// TIA Portal project "Motor with VFD+PID" (V20)

(* hardware
DEVICE "S7-1200 station_1"  S7-1200 Station
   slot 0: "Rack_0"  S7-1200 Rack  Rack  V1.0
   slot 1: "PLC_1"  CPU 1214C DC/DC/DC  6ES7 214-1AG40-0XB0  V4.7
DEVICE "HMI_1"  KTP700 Basic PN
   slot 0: "HMI_1"  KTP700 Basic PN  6AV2 123-2GB03-0AX0  17.0.0.0
   slot 1: "HMI_RT_1"  KTP700 Basic PN  6AV2 123-2GB03-0AX0  17.0.0.0
   slot 5: "HMI_1.IE_CP_1"  PROFINET Interface  17.0.0.0
      slot 1: "PROFINET Interface_1"  PROFINET Interface
         slot 1: "Port_1"  Port
*)

// ===== PLC "PLC_1"  CPU 1214C DC/DC/DC =====

VAR_GLOBAL   // PLC tag table "Default tag table"
   "Start_PB" AT %I0.0 : Bool;
   "Stop_PB" AT %I0.1 : Bool;
   "VFD_Fault" AT %I0.2 : Bool;
   "VFD_Running_FB" AT %I0.3 : Bool;
   "Reset_PB" AT %I0.4 : Bool;
   "VFD_Run_CMD" AT %Q0.0 : Bool;
   "VFD_Reset_CMD" AT %Q0.1 : Bool;
   "Motor_Run_Latch" AT %M0.0 : Bool;
   "Alarm_Active" AT %M0.1 : Bool;
   "Auto_Mode" AT %M0.2 : Bool;
   "Manual_Mode" AT %M0.3 : Bool;
   "HMI_START" AT %M0.4 : Bool;
   "HMI_STOP" AT %M0.5 : Bool;
   "HMI_RESET" AT %M0.6 : Bool;
END_VAR

DATA_BLOCK "DB_VFD_Motor"   // DB1
{ S7_Optimized_Access := 'TRUE' }
VERSION : 0.1
   VAR RETAIN
      Speed_setpoint_hz : Real := 25.0;
   END_VAR
   VAR
      Max_Hz : Real := 50.0;
      Min_Hz : Real;
      Pressure_Setpoint : Real := 6.0;
      Ramp_Output : Real;
      Ramp_Step : Real := 1.0;
      Pressure_Actual : Real := 4.0;
      PID_Error : Real;
   END_VAR
   VAR RETAIN
      Ramp_time : Real;
   END_VAR
   VAR
      Low_Pressure_timer_Done : Bool;
      Min_Pressure_Limit : Real := 1.0;
      Max_Pressure_Limit : Real := 8.0;
      Manual_Speed_Hz : Real := 20.0;
      Overpressure_Alarm : Bool;
      Low_Pressure_Alarm : Bool;
      Fault_code : Int;
      Actual_speed_hz : Real;
      Output_scaled : Int;
   END_VAR
BEGIN
END_DATA_BLOCK

// folder: System blocks/Program resources

DATA_BLOCK "TON"   // DB2
{ S7_Optimized_Access := 'TRUE' }
AUTHOR : Simatic
FAMILY : IEC
NAME : IEC_TMR
VERSION : 1.0
// stored: InstanceOfName IEC_TIMER
"IEC_TIMER"
BEGIN
END_DATA_BLOCK

// folder: (top level)

ORGANIZATION_BLOCK "Main"   // OB1, LAD, ProgramCycle
TITLE = "Main Program Sweep (Cycle)"
{ S7_Optimized_Access := 'TRUE' }
VERSION : 0.1
   VAR_INPUT
      Initial_Call : Bool;   // Initial call of this OB
      Remanence : Bool;   // =True, if remanent data are available
   END_VAR
BEGIN

REGION Network 1: Start/Stop Safety Logic
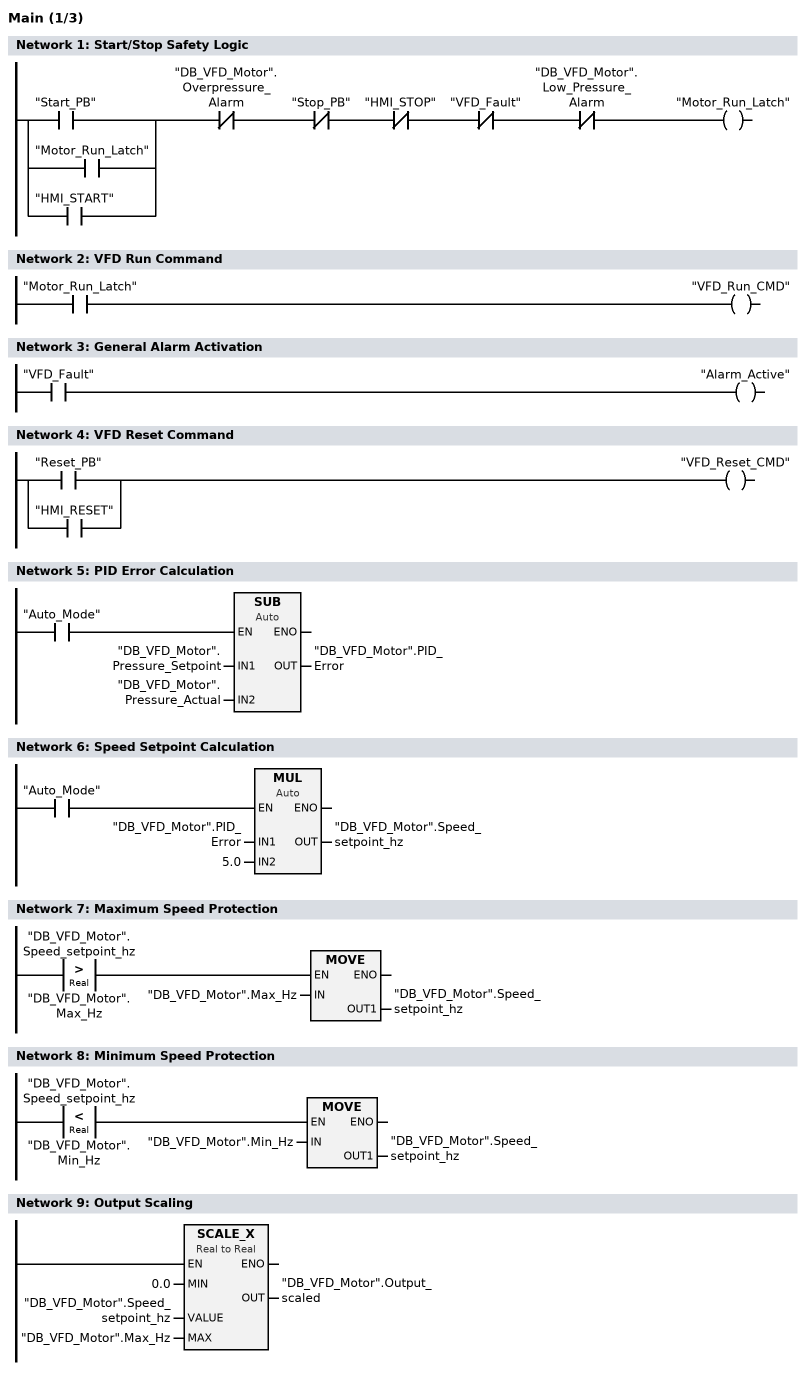
   RUNG wire#powerrail
      Contact( "Start_PB" )
      wire#w1
      I_Contact( "DB_VFD_Motor".Overpressure_Alarm )
      I_Contact( "Stop_PB" )
      I_Contact( "HMI_STOP" )
      I_Contact( "VFD_Fault" )
      I_Contact( "DB_VFD_Motor".Low_Pressure_Alarm )
      Coil( "Motor_Run_Latch" )
   END_RUNG
   RUNG wire#powerrail
      Contact( "Motor_Run_Latch" )
   END_RUNG wire#w1
   RUNG wire#powerrail
      Contact( "HMI_START" )
   END_RUNG wire#w1
   // the same network as SCL:
   "Motor_Run_Latch" := ("Start_PB" OR "Motor_Run_Latch" OR "HMI_START") AND NOT "DB_VFD_Motor".Overpressure_Alarm AND NOT "Stop_PB" AND NOT "HMI_STOP" AND NOT "VFD_Fault" AND NOT "DB_VFD_Motor".Low_Pressure_Alarm;
END_REGION

REGION Network 2: VFD Run Command
   RUNG wire#powerrail
      Contact( "Motor_Run_Latch" )
      Coil( "VFD_Run_CMD" )
   END_RUNG
   // the same network as SCL:
   "VFD_Run_CMD" := "Motor_Run_Latch";
END_REGION

REGION Network 3: General Alarm Activation
   RUNG wire#powerrail
      Contact( "VFD_Fault" )
      Coil( "Alarm_Active" )
   END_RUNG
   // the same network as SCL:
   "Alarm_Active" := "VFD_Fault";
END_REGION

REGION Network 4: VFD Reset Command
   RUNG wire#powerrail
      Contact( "Reset_PB" )
      wire#w1
      Coil( "VFD_Reset_CMD" )
   END_RUNG
   RUNG wire#powerrail
      Contact( "HMI_RESET" )
   END_RUNG wire#w1
   // the same network as SCL:
   "VFD_Reset_CMD" := "Reset_PB" OR "HMI_RESET";
END_REGION

REGION Network 5: PID Error Calculation
   RUNG wire#powerrail
      Contact( "Auto_Mode" )
      Sub(in1 := "DB_VFD_Motor".Pressure_Setpoint, in2 := "DB_VFD_Motor".Pressure_Actual, out => "DB_VFD_Motor".PID_Error)
   END_RUNG
   // the same network as SCL:
   IF "Auto_Mode" THEN
       "DB_VFD_Motor".PID_Error := "DB_VFD_Motor".Pressure_Setpoint - "DB_VFD_Motor".Pressure_Actual;
   END_IF;
END_REGION

REGION Network 6: Speed Setpoint Calculation
   RUNG wire#powerrail
      Contact( "Auto_Mode" )
      Mul(in1 := "DB_VFD_Motor".PID_Error, in2 := 5.0, out => "DB_VFD_Motor".Speed_setpoint_hz)
   END_RUNG
   // the same network as SCL:
   IF "Auto_Mode" THEN "DB_VFD_Motor".Speed_setpoint_hz := "DB_VFD_Motor".PID_Error * 5.0; END_IF;
END_REGION

REGION Network 7: Maximum Speed Protection
   RUNG wire#powerrail
      { S7_Templates := "SrcType := Real" } GT_Contact(in1 := "DB_VFD_Motor".Speed_setpoint_hz, in2 := "DB_VFD_Motor".Max_Hz)
      Move(in := "DB_VFD_Motor".Max_Hz, out1 => "DB_VFD_Motor".Speed_setpoint_hz)
   END_RUNG
   // the same network as SCL:
   IF "DB_VFD_Motor".Speed_setpoint_hz > "DB_VFD_Motor".Max_Hz THEN
       "DB_VFD_Motor".Speed_setpoint_hz := "DB_VFD_Motor".Max_Hz;
   END_IF;
END_REGION

REGION Network 8: Minimum Speed Protection
   RUNG wire#powerrail
      { S7_Templates := "SrcType := Real" } LT_Contact(in1 := "DB_VFD_Motor".Speed_setpoint_hz, in2 := "DB_VFD_Motor".Min_Hz)
      Move(in := "DB_VFD_Motor".Min_Hz, out1 => "DB_VFD_Motor".Speed_setpoint_hz)
   END_RUNG
   // the same network as SCL:
   IF "DB_VFD_Motor".Speed_setpoint_hz < "DB_VFD_Motor".Min_Hz THEN
       "DB_VFD_Motor".Speed_setpoint_hz := "DB_VFD_Motor".Min_Hz;
   END_IF;
END_REGION

REGION Network 9: Output Scaling
   RUNG wire#powerrail
      { S7_Templates := "[SrcType := Real, DestType := Real]" } Scale(min := 0.0, value := "DB_VFD_Motor".Speed_setpoint_hz, max := "DB_VFD_Motor".Max_Hz, out => "DB_VFD_Motor".Output_scaled)
   END_RUNG
   // the same network as SCL:
   "DB_VFD_Motor".Output_scaled := SCALE_X(MIN := 0.0, VALUE := "DB_VFD_Motor".Speed_setpoint_hz, MAX := "DB_VFD_Motor".Max_Hz);
END_REGION

REGION Network 10: Motor Speed Update
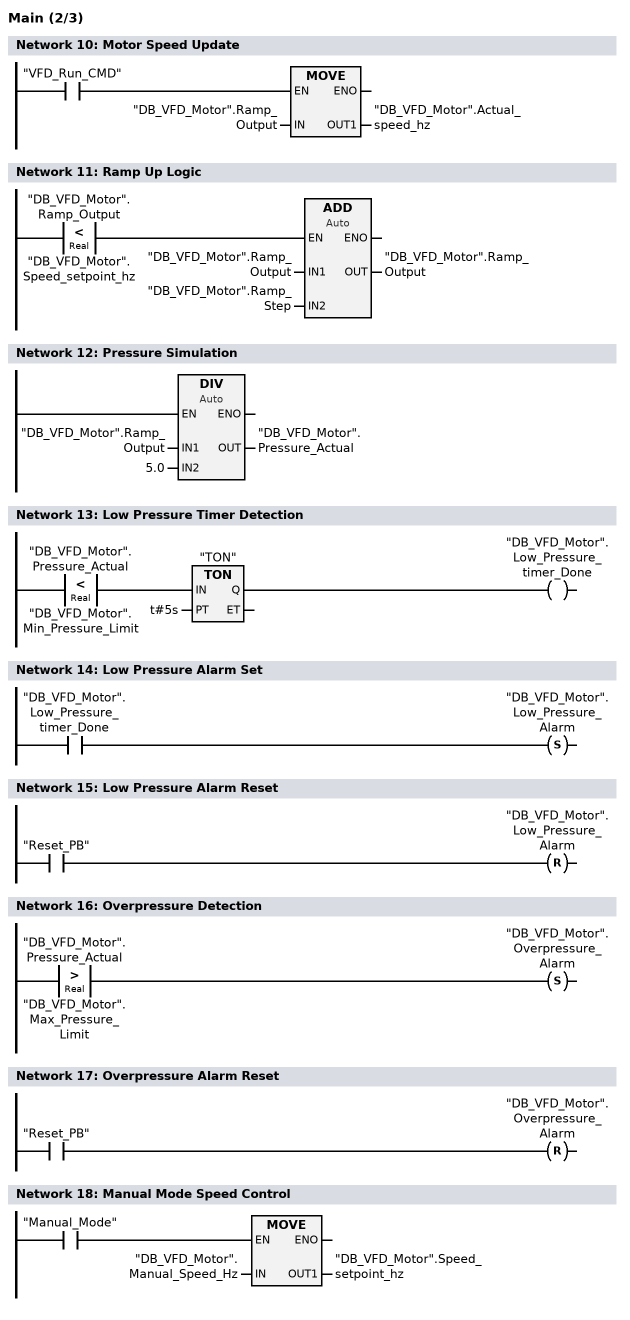
   RUNG wire#powerrail
      Contact( "VFD_Run_CMD" )
      Move(in := "DB_VFD_Motor".Ramp_Output, out1 => "DB_VFD_Motor".Actual_speed_hz)
   END_RUNG
   // the same network as SCL:
   IF "VFD_Run_CMD" THEN "DB_VFD_Motor".Actual_speed_hz := "DB_VFD_Motor".Ramp_Output; END_IF;
END_REGION

REGION Network 11: Ramp Up Logic
   RUNG wire#powerrail
      { S7_Templates := "SrcType := Real" } LT_Contact(in1 := "DB_VFD_Motor".Ramp_Output, in2 := "DB_VFD_Motor".Speed_setpoint_hz)
      Add(in1 := "DB_VFD_Motor".Ramp_Output, in2 := "DB_VFD_Motor".Ramp_Step, out => "DB_VFD_Motor".Ramp_Output)
   END_RUNG
   // the same network as SCL:
   IF "DB_VFD_Motor".Ramp_Output < "DB_VFD_Motor".Speed_setpoint_hz THEN
       "DB_VFD_Motor".Ramp_Output := "DB_VFD_Motor".Ramp_Output + "DB_VFD_Motor".Ramp_Step;
   END_IF;
END_REGION

REGION Network 12: Pressure Simulation
   RUNG wire#powerrail
      Div(in1 := "DB_VFD_Motor".Ramp_Output, in2 := 5.0, out => "DB_VFD_Motor".Pressure_Actual)
   END_RUNG
   // the same network as SCL:
   "DB_VFD_Motor".Pressure_Actual := "DB_VFD_Motor".Ramp_Output / 5.0;
END_REGION

REGION Network 13: Low Pressure Timer Detection
   "TON".TON(IN := "DB_VFD_Motor".Pressure_Actual < "DB_VFD_Motor".Min_Pressure_Limit, PT := t#5s);
   "DB_VFD_Motor".Low_Pressure_timer_Done := "TON".Q;
END_REGION

REGION Network 14: Low Pressure Alarm Set
   RUNG wire#powerrail
      Contact( "DB_VFD_Motor".Low_Pressure_timer_Done )
      S_Coil( "DB_VFD_Motor".Low_Pressure_Alarm )
   END_RUNG
   // the same network as SCL:
   IF "DB_VFD_Motor".Low_Pressure_timer_Done THEN "DB_VFD_Motor".Low_Pressure_Alarm := TRUE; END_IF;
END_REGION

REGION Network 15: Low Pressure Alarm Reset
   RUNG wire#powerrail
      Contact( "Reset_PB" )
      R_Coil( "DB_VFD_Motor".Low_Pressure_Alarm )
   END_RUNG
   // the same network as SCL:
   IF "Reset_PB" THEN "DB_VFD_Motor".Low_Pressure_Alarm := FALSE; END_IF;
END_REGION

REGION Network 16: Overpressure Detection
   RUNG wire#powerrail
      { S7_Templates := "SrcType := Real" } GT_Contact(in1 := "DB_VFD_Motor".Pressure_Actual, in2 := "DB_VFD_Motor".Max_Pressure_Limit)
      S_Coil( "DB_VFD_Motor".Overpressure_Alarm )
   END_RUNG
   // the same network as SCL:
   IF "DB_VFD_Motor".Pressure_Actual > "DB_VFD_Motor".Max_Pressure_Limit THEN
       "DB_VFD_Motor".Overpressure_Alarm := TRUE;
   END_IF;
END_REGION

REGION Network 17: Overpressure Alarm Reset
   RUNG wire#powerrail
      Contact( "Reset_PB" )
      R_Coil( "DB_VFD_Motor".Overpressure_Alarm )
   END_RUNG
   // the same network as SCL:
   IF "Reset_PB" THEN "DB_VFD_Motor".Overpressure_Alarm := FALSE; END_IF;
END_REGION

REGION Network 18: Manual Mode Speed Control
   RUNG wire#powerrail
      Contact( "Manual_Mode" )
      Move(in := "DB_VFD_Motor".Manual_Speed_Hz, out1 => "DB_VFD_Motor".Speed_setpoint_hz)
   END_RUNG
   // the same network as SCL:
   IF "Manual_Mode" THEN "DB_VFD_Motor".Speed_setpoint_hz := "DB_VFD_Motor".Manual_Speed_Hz; END_IF;
END_REGION

REGION Network 19: VFD Fault Code Assignment
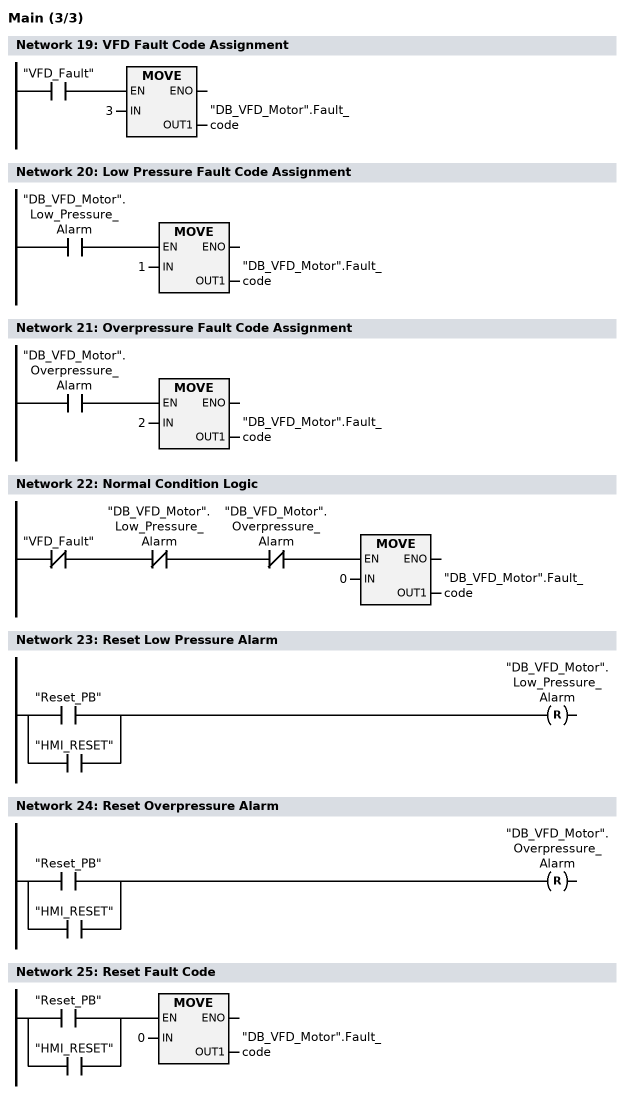
   RUNG wire#powerrail
      Contact( "VFD_Fault" )
      Move(in := 3, out1 => "DB_VFD_Motor".Fault_code)
   END_RUNG
   // the same network as SCL:
   IF "VFD_Fault" THEN "DB_VFD_Motor".Fault_code := 3; END_IF;
END_REGION

REGION Network 20: Low Pressure Fault Code Assignment
   RUNG wire#powerrail
      Contact( "DB_VFD_Motor".Low_Pressure_Alarm )
      Move(in := 1, out1 => "DB_VFD_Motor".Fault_code)
   END_RUNG
   // the same network as SCL:
   IF "DB_VFD_Motor".Low_Pressure_Alarm THEN "DB_VFD_Motor".Fault_code := 1; END_IF;
END_REGION

REGION Network 21: Overpressure Fault Code Assignment
   RUNG wire#powerrail
      Contact( "DB_VFD_Motor".Overpressure_Alarm )
      Move(in := 2, out1 => "DB_VFD_Motor".Fault_code)
   END_RUNG
   // the same network as SCL:
   IF "DB_VFD_Motor".Overpressure_Alarm THEN "DB_VFD_Motor".Fault_code := 2; END_IF;
END_REGION

REGION Network 22: Normal Condition Logic
   RUNG wire#powerrail
      I_Contact( "VFD_Fault" )
      I_Contact( "DB_VFD_Motor".Low_Pressure_Alarm )
      I_Contact( "DB_VFD_Motor".Overpressure_Alarm )
      Move(in := 0, out1 => "DB_VFD_Motor".Fault_code)
   END_RUNG
   // the same network as SCL:
   IF NOT "VFD_Fault" AND NOT "DB_VFD_Motor".Low_Pressure_Alarm AND NOT "DB_VFD_Motor".Overpressure_Alarm THEN
       "DB_VFD_Motor".Fault_code := 0;
   END_IF;
END_REGION

REGION Network 23: Reset Low Pressure Alarm
   RUNG wire#powerrail
      Contact( "Reset_PB" )
      wire#w1
      R_Coil( "DB_VFD_Motor".Low_Pressure_Alarm )
   END_RUNG
   RUNG wire#powerrail
      Contact( "HMI_RESET" )
   END_RUNG wire#w1
   // the same network as SCL:
   IF "Reset_PB" OR "HMI_RESET" THEN "DB_VFD_Motor".Low_Pressure_Alarm := FALSE; END_IF;
END_REGION

REGION Network 24: Reset Overpressure Alarm
   RUNG wire#powerrail
      Contact( "Reset_PB" )
      wire#w1
      R_Coil( "DB_VFD_Motor".Overpressure_Alarm )
   END_RUNG
   RUNG wire#powerrail
      Contact( "HMI_RESET" )
   END_RUNG wire#w1
   // the same network as SCL:
   IF "Reset_PB" OR "HMI_RESET" THEN "DB_VFD_Motor".Overpressure_Alarm := FALSE; END_IF;
END_REGION

REGION Network 25: Reset Fault Code
   RUNG wire#powerrail
      Contact( "Reset_PB" )
      wire#w1
      Move(in := 0, out1 => "DB_VFD_Motor".Fault_code)
   END_RUNG
   RUNG wire#powerrail
      Contact( "HMI_RESET" )
   END_RUNG wire#w1
   // the same network as SCL:
   IF "Reset_PB" OR "HMI_RESET" THEN "DB_VFD_Motor".Fault_code := 0; END_IF;
END_REGION
END_ORGANIZATION_BLOCK

(* ===== HMI "HMI_RT_1" =====
system functions are stored by id; their names below are inferred from use
connection "HMI_Connection_1": ETHERNET, SMART_S7_1200_OMS

HMI tags "Default tag table"
   "Tag_ScreenNumber" : UInt, internal
   "Motor_Run_Latch" : Bool = PLC Motor_Run_Latch AT %M0.0, 1 s
   "Alarm_Active" : Bool = PLC Alarm_Active AT %M0.1, 1 s
   "Auto_Mode" : Bool = PLC Auto_Mode AT %M0.2, 1 s
   "Manual_Mode" : Bool = PLC Manual_Mode AT %M0.3, 1 s
   "HMI_START" : Bool = PLC HMI_START AT %M0.4, 1 s
   "HMI_STOP" : Bool = PLC HMI_STOP AT %M0.5, 1 s
   "HMI_RESET" : Bool = PLC HMI_RESET AT %M0.6, 1 s
   "DB_VFD_Motor_Pressure_Setpoint" : Real = PLC DB_VFD_Motor.Pressure_Setpoint, 1 s
   "DB_VFD_Motor_Pressure_Actual" : Real = PLC DB_VFD_Motor.Pressure_Actual, 1 s
   "DB_VFD_Motor_Actual_speed_hz" : Real = PLC DB_VFD_Motor.Actual_speed_hz, 1 s
   "DB_VFD_Motor_Output_scaled" : Int = PLC DB_VFD_Motor.Output_scaled, 1 s
   "DB_VFD_Motor_Manual_Speed_Hz" : Real = PLC DB_VFD_Motor.Manual_Speed_Hz, 1 s
   "DB_VFD_Motor_PID_Error" : Real = PLC DB_VFD_Motor.PID_Error, 1 s
   "DB_VFD_Motor_Speed_setpoint_hz" : Real = PLC DB_VFD_Motor.Speed_setpoint_hz, 1 s
   "DB_VFD_Motor_Ramp_Output" : Real = PLC DB_VFD_Motor.Ramp_Output, 1 s
   "DB_VFD_Motor_Min_Pressure_Limit" : Real = PLC DB_VFD_Motor.Min_Pressure_Limit, 1 s
   "DB_VFD_Motor_Max_Pressure_Limit" : Real = PLC DB_VFD_Motor.Max_Pressure_Limit, 1 s
   "DB_VFD_Motor_Ramp_Step" : Real = PLC DB_VFD_Motor.Ramp_Step, 1 s
   "DB_VFD_Motor_Fault_code" : Int = PLC DB_VFD_Motor.Fault_code, 1 s
   "VFD_Fault" : Bool = PLC VFD_Fault AT %I0.2, 1 s
   "DB_VFD_Motor_Low_Pressure_Alarm" : Bool = PLC DB_VFD_Motor.Low_Pressure_Alarm, 1 s
   "DB_VFD_Motor_Overpressure_Alarm" : Bool = PLC DB_VFD_Motor.Overpressure_Alarm, 1 s

text list "ACTIVE": 0 'INACTIVE'; 1 'ACTIVE'

text list "RUNNING": 0 'STOPPED'; 1 'RUNNING'

text list "ALARM": 0 'NO ALARM'; 1 'ALARM'

text list "NO FAULT": 0 'NO FAULT'; 1 'VFD FAULT ACTIVE'

text list "NO ALARM": 0 'NO ALARM'; 1 'LOW PRESSURE ACTIVE'

text list "OVERPRESSURE ACTIVE": 0 'NO ALARM'; 1 'OVERPRESSURE ACTIVE'

Template "Template_1" 800x480
   Button "Exit" at 714,429 size 71x50; TextOff 'Exit'; PictureOff "ExitRuntime_KTP700_Basic_PN_TR"; PictureOn "ExitRuntime_KTP700_Basic_PN_TR"
      on Release: StopRuntime(0)
   Button "Template_Button" at 614,429 size 71x50; TextOff 'Text'
   Button "Template_Button_1" at 514,429 size 71x50; TextOff 'Text'
   Button "Template_Button_2" at 414,429 size 71x50; TextOff 'Text'
   Button "Template_Button_3" at 314,429 size 71x50; TextOff 'Text'
   Button "Template_Button_4" at 214,429 size 71x50; TextOff 'Text'
   Button "Template_Button_5" at 114,429 size 71x50; TextOff 'Text'
   Button "Start screen" at 14,429 size 71x50; TextOff 'Start screen'; PictureOff "NavigateHome_KTP700_Basic_PN_TR"; PictureOn "NavigateHome_KTP700_Basic_PN_TR"
      on Release: ActivateScreen("Main Overview", 0)
   SymbolicIOField "Symbolic_IO_Field_Screen" at 93,9 size 600x33; TextOff '0'; TextOn '1'; TextList "TextList_ScreenNames"
      ProcessValue <- "Tag_ScreenNumber"
      on Change: ActivateScreenByNumber("Tag_ScreenNumber", 0)
   DateTimeField "HmiScreenItemData" at 695,25 size 105x25
   DateTimeField "HmiScreenItemData_1" at 695,0 size 105x25
   GraphicView "Logo" at 0,0 size 91x51; Picture "Logo of HMI_1"

screen "Main Overview" 800x480, template "Template_1"
   on GenerateScreen: SetTag("Tag_ScreenNumber", 1)
   GraphicView "Graphic view_1" at 2,1 size 796x478; Picture "ChatGPT Image 23 Ιουν 2026, 10_41_49 μ.μ."
   TextField "Text field_1" at 235,6 size 313x27; Text 'VFD PUMP PRESSURE CONTROL'
   GraphicView "Graphic view_2" at 123,75 size 264x225; Picture "ChatGPT Image 23 Ιουν 2026, 10_44_50 μ.μ."
   TextField "Text field_2" at 304,43 size 150x25; Text 'MAIN OVERVIEW'
   Button "Button_1" at 146,332 size 144x62; TextOff 'START'
      on Press: function_b14e0dd5("HMI_START", 0)
   Button "Button_2" at 1,414 size 194x65; TextOff 'HOME'
   Button "Button_3" at 195,414 size 204x65; TextOff 'CONTROL'
      on Press: ActivateScreen("Control", 0)
   Button "Button_4" at 398,414 size 200x65; TextOff 'ALARMS'
      on Press: ActivateScreen("Alarm Page", 0)
   Button "Button_5" at 597,414 size 200x65; TextOff 'DIAGNOSTICS'
      on Press: ActivateScreen("Diagnostics", 0)
   Button "Button_6" at 304,332 size 144x62; TextOff 'STOP'
      on Press: function_b14e0dd5("HMI_STOP", 0)
   Button "Button_7" at 462,332 size 144x62; TextOff 'RESET'
      on Press: function_b14e0dd5("HMI_RESET", 0)
   GraphicView "Graphic view_3" at 385,87 size 192x28; Picture "ChatGPT Image 23 Ιουν 2026, 10_41_49 μ.μ._2"
   GraphicView "Graphic view_4" at 594,87 size 192x28; Picture "ChatGPT Image 23 Ιουν 2026, 10_41_49 μ.μ._2"
   GraphicView "Graphic view_6" at 385,200 size 129x35; Picture "ChatGPT Image 23 Ιουν 2026, 10_41_49 μ.μ._2"
   IOField "I/O field_2" at 628,124 size 122x53; FormatPattern 99.9; Unit bar
      ProcessValue <- "DB_VFD_Motor_Pressure_Actual"
   IOField "I/O field_3" at 389,242 size 122x53; FormatPattern 99.9; Unit Hz
      ProcessValue <- "DB_VFD_Motor_Manual_Speed_Hz"
   GraphicView "Graphic view_7" at 610,430 size 39x34; Picture "Graphic_1"
   GraphicView "Graphic view_8" at 422,429 size 43x33; Picture "Graphic_2"
   GraphicView "Graphic view_9" at 35,428 size 41x33; Picture "Graphic_3"
   GraphicView "Graphic view_10" at 213,430 size 36x30; Picture "Graphic_4"
   Circle "Circle_1" at 13,86 size 29x29
      Appearance <- "Motor_Run_Latch"
   Circle "Circle_2" at 13,137 size 29x29
      Appearance <- "Alarm_Active"
   Circle "Circle_3" at 13,185 size 29x29
      Appearance <- "Auto_Mode"
   Circle "Circle_4" at 13,235 size 29x29
      Appearance <- "Manual_Mode"
   TextField "Text field_3" at 46,84 size 102x20; Text 'MOTOR STATUS'
   TextField "Text field_4" at 44,137 size 104x20; Text 'ALARM STATUS'
   TextField "Text field_5" at 47,182 size 79x20; Text 'AUTO MODE'
   TextField "Text field_6" at 46,233 size 99x20; Text 'MANUAL MODE'
   SymbolicIOField "Symbolic I/O field_1" at 45,253 size 75x25; TextOff '0'; TextOn '1'; TextList "ACTIVE"
      ProcessValue <- "Manual_Mode"
      Appearance <- "Manual_Mode"
   SymbolicIOField "Symbolic I/O field_2" at 47,204 size 75x25; TextOff '0'; TextOn '1'; TextList "ACTIVE"
      ProcessValue <- "Auto_Mode"
      Appearance <- "Auto_Mode"
   SymbolicIOField "Symbolic I/O field_3" at 46,103 size 77x20; TextOff '0'; TextOn '1'; TextList "RUNNING"
      ProcessValue <- "Motor_Run_Latch"
      Appearance <- "Motor_Run_Latch"
   SymbolicIOField "Symbolic I/O field_4" at 46,157 size 83x18; TextOff '0'; TextOn '1'; TextList "ALARM"
      ProcessValue <- "Alarm_Active"
      Appearance <- "Alarm_Active"
   TextField "Text field_7" at 418,92 size 132x20; Text 'PRESSURE SETPOINT'
   TextField "Text field_8" at 620,91 size 136x20; Text 'ACTUAL PRESSPOINT'
   TextField "Text field_9" at 401,201 size 106x36; Text 'MANUAL SPEED SETPOINT'
   IOField "I/O field_1" at 412,124 size 122x53; FormatPattern 99.9; Unit bar
      ProcessValue <- "DB_VFD_Motor_Pressure_Setpoint"
   GraphicView "Graphic view_5" at 522,201 size 129x35; Picture "ChatGPT Image 23 Ιουν 2026, 10_41_49 μ.μ._2"
   TextField "Text field_11" at 538,199 size 108x36; Text 'ACTUAL MOTOR SPEED'
   IOField "I/O field_5" at 522,243 size 127x53; FormatPattern 99.99; Unit Hz
      ProcessValue <- "DB_VFD_Motor_Actual_speed_hz"
   GraphicView "Graphic view_11" at 657,200 size 129x35; Picture "ChatGPT Image 23 Ιουν 2026, 10_41_49 μ.μ._2"
   TextField "Text field_10" at 672,205 size 105x20; Text 'OUTPUT SCALED'
   IOField "I/O field_4" at 662,245 size 122x53; FormatPattern 9999; Unit %
      ProcessValue <- "DB_VFD_Motor_Output_scaled"

screen "Control" 800x480, template "Template_1"
   on GenerateScreen: SetTag("Tag_ScreenNumber", 1)
   GraphicView "Graphic view_1" at 2,1 size 796x478; Picture "ChatGPT Image 23 Ιουν 2026, 10_41_49 μ.μ."
   TextField "Text field_1" at 235,6 size 313x27; Text 'VFD PUMP PRESSURE CONTROL'
   TextField "Text field_2" at 351,42 size 87x25; Text 'CONTROL'
   Button "Button_2" at 1,414 size 194x65; TextOff 'HOME'
      on Press: ActivateScreen("Main Overview", 0)
   Button "Button_3" at 195,414 size 204x65; TextOff 'CONTROL'
      on Press: ActivateScreen("Control", 0)
   Button "Button_4" at 398,414 size 200x65; TextOff 'ALARMS'
      on Press: ActivateScreen("Alarm Page", 0)
   Button "Button_5" at 597,414 size 200x65; TextOff 'DIAGNOSTICS'
      on Press: ActivateScreen("Diagnostics", 0)
   GraphicView "Graphic view_4" at 472,128 size 304x28; Picture "ChatGPT Image 23 Ιουν 2026, 10_41_49 μ.μ._2"
   GraphicView "Graphic view_7" at 610,430 size 39x34; Picture "Graphic_1"
   GraphicView "Graphic view_8" at 422,429 size 43x33; Picture "Graphic_2"
   GraphicView "Graphic view_9" at 35,428 size 41x33; Picture "Graphic_3"
   GraphicView "Graphic view_10" at 213,430 size 36x30; Picture "Graphic_4"
   TextField "Text field_4" at 27,92 size 111x20; Text 'MODE SELECTION'
   TextField "Text field_5" at 235,136 size 79x20; Text 'AUTO MODE'
   TextField "Text field_6" at 228,226 size 99x20; Text 'MANUAL MODE'
   Button "Button_7" at 17,209 size 144x74; TextOff 'MANUAL MODE'
      on Activate: SetBit("Manual_Mode"); ResetBit("Auto_Mode")
   Button "Button_1" at 17,128 size 144x72; TextOff 'AUTO MODE'
      on Activate: SetBit("Auto_Mode"); ResetBit("Manual_Mode")
   GraphicView "Graphic view_2" at 471,235 size 304x28; Picture "ChatGPT Image 23 Ιουν 2026, 10_41_49 μ.μ._2"
   GraphicView "Graphic view_3" at 407,337 size 163x28; Picture "ChatGPT Image 23 Ιουν 2026, 10_41_49 μ.μ._2"
   GraphicView "Graphic view_5" at 214,337 size 163x28; Picture "ChatGPT Image 23 Ιουν 2026, 10_41_49 μ.μ._2"
   GraphicView "Graphic view_6" at 25,337 size 155x28; Picture "ChatGPT Image 23 Ιουν 2026, 10_41_49 μ.μ._2"
   GraphicView "Graphic view_11" at 603,338 size 163x28; Picture "ChatGPT Image 23 Ιουν 2026, 10_41_49 μ.μ._2"
   SymbolicIOField "Symbolic I/O field_2" at 236,155 size 75x25; TextOff '0'; TextOn '1'; TextList "ACTIVE"
      ProcessValue <- "Auto_Mode"
      Appearance <- "Auto_Mode"
   SymbolicIOField "Symbolic I/O field_1" at 231,246 size 75x25; TextOff '0'; TextOn '1'; TextList "ACTIVE"
      ProcessValue <- "Manual_Mode"
      Appearance <- "Manual_Mode"
   Circle "Circle_1" at 199,141 size 29x29
      Appearance <- "Auto_Mode"
   Circle "Circle_4" at 199,231 size 29x29
      Appearance <- "Manual_Mode"
   IOField "I/O field_2" at 569,157 size 142x53; FormatPattern 99.9; Unit bar
      ProcessValue <- "DB_VFD_Motor_Pressure_Setpoint"
   TextField "Text field_7" at 563,132 size 132x20; Text 'PRESSURE SETPOINT'
   IOField "I/O field_3" at 567,267 size 115x53; FormatPattern 99.9; Unit Hz
      ProcessValue <- "DB_VFD_Motor_Manual_Speed_Hz"
   TextField "Text field_9" at 548,239 size 165x20; Text 'MANUAL SPEED SETPOINT'
   TextField "Text field_3" at 61,340 size 74x20; Text 'PID ERROR'
   TextField "Text field_8" at 238,341 size 111x20; Text 'SPEED SETPOINT'
   TextField "Text field_10" at 438,341 size 94x20; Text 'RAMP OUTPUT'
   TextField "Text field_11" at 633,342 size 98x20; Text 'ACTUAL SPEED'
   IOField "I/O field_1" at 231,366 size 134x40; FormatPattern 99.9; Unit Hz
      ProcessValue <- "DB_VFD_Motor_Speed_setpoint_hz"
   IOField "I/O field_4" at 426,368 size 134x40; FormatPattern 99.9; Unit Hz
      ProcessValue <- "DB_VFD_Motor_Ramp_Output"
   IOField "I/O field_5" at 620,369 size 134x40; FormatPattern 99.9; Unit Hz
      ProcessValue <- "DB_VFD_Motor_Actual_speed_hz"
   IOField "I/O field_6" at 24,370 size 154x37; FormatPattern 99.9; Unit bar
      ProcessValue <- "DB_VFD_Motor_PID_Error"

screen "Alarm Page" 800x480, template "Template_1"
   on GenerateScreen: SetTag("Tag_ScreenNumber", 1)
   GraphicView "Graphic view_1" at 0,1 size 799x478; Picture "ChatGPT Image 23 Ιουν 2026, 10_41_49 μ.μ."
   TextField "Text field_1" at 235,6 size 313x27; Text 'VFD PUMP PRESSURE CONTROL'
   TextField "Text field_2" at 352,38 size 77x25; Text 'ALARMS'
   Button "Button_2" at 1,414 size 194x65; TextOff 'HOME'
      on Press: ActivateScreen("Main Overview", 0)
   Button "Button_3" at 195,414 size 204x65; TextOff 'CONTROL'
      on Press: ActivateScreen("Control", 0)
   Button "Button_4" at 398,414 size 200x65; TextOff 'ALARMS'
      on Press: ActivateScreen("Alarm Page", 0)
   Button "Button_5" at 597,414 size 200x65; TextOff 'DIAGNOSTICS'
      on Press: ActivateScreen("Diagnostics", 0)
   GraphicView "Graphic view_7" at 610,430 size 39x34; Picture "Graphic_1"
   GraphicView "Graphic view_8" at 422,429 size 43x33; Picture "Graphic_2"
   GraphicView "Graphic view_9" at 35,428 size 41x33; Picture "Graphic_3"
   GraphicView "Graphic view_10" at 213,430 size 36x30; Picture "Graphic_4"
   Circle "Circle_4" at 249,194 size 29x29
      Appearance <- "DB_VFD_Motor_Low_Pressure_Alarm"
   TextField "Text field_3" at 25,337 size 80x20; Text 'FAULT CODE'
   TextField "Text field_4" at 58,96 size 56x20; Text 'ALARM'
   TextField "Text field_5" at 21,251 size 154x20; Text 'OVERPRESSURE ALARM'
   TextField "Text field_6" at 40,138 size 71x20; Text 'VFD FAULT'
   Circle "Circle_1" at 249,135 size 29x29
      Appearance <- "VFD_Fault"
   TextField "Text field_7" at 240,98 size 53x20; Text 'STATUS'
   Circle "Circle_2" at 249,269 size 29x29
      Appearance <- "DB_VFD_Motor_Overpressure_Alarm"
   TextField "Text field_8" at 391,100 size 88x20; Text 'DESCRIPTION'
   IOField "I/O field_1" at 330,340 size 17x32; FormatPattern 9
      ProcessValue <- "DB_VFD_Motor_Fault_code"
   TextField "Text field_9" at 599,93 size 98x20; Text 'ALARM RESET'
   TextField "Text field_10" at 592,215 size 130x20; Text 'FAULT CODE LEGEND'
   TextField "Text field_11" at 544,255 size 110x23; Text '0=NO FAULT'
   TextField "Text field_12" at 543,282 size 157x23; Text '1=LOW PRESSURE'
   TextField "Text field_13" at 542,310 size 160x23; Text '2=OVERPRESSURE'
   TextField "Text field_14" at 542,340 size 118x23; Text '3=VFD FAULT'
   TextField "Text field_15" at 22,174 size 153x20; Text 'LOW PRESSURE ALARM'
   SymbolicIOField "Symbolic I/O field_1" at 349,136 size 102x23; TextOff '0'; TextOn '1'; TextList "NO FAULT"
      ProcessValue <- "VFD_Fault"
      Appearance <- "VFD_Fault"
   SymbolicIOField "Symbolic I/O field_2" at 340,189 size 162x39; TextOff '0'; TextOn '1'; TextList "NO ALARM"
      Appearance <- "DB_VFD_Motor_Low_Pressure_Alarm"
      ProcessValue <- "DB_VFD_Motor_Low_Pressure_Alarm"
   SymbolicIOField "Symbolic I/O field_3" at 342,266 size 160x40; TextOff '0'; TextOn '1'; TextList "OVERPRESSURE ACTIVE"
      ProcessValue <- "DB_VFD_Motor_Overpressure_Alarm"
      Appearance <- "DB_VFD_Motor_Overpressure_Alarm"
   Button "Button_7" at 553,127 size 187x62; TextOff 'RESET'
      on Press: function_b14e0dd5("HMI_RESET", 0)

screen "Diagnostics" 800x480, template "Template_1"
   on GenerateScreen: SetTag("Tag_ScreenNumber", 1)
   GraphicView "Graphic view_1" at 2,1 size 796x478; Picture "ChatGPT Image 23 Ιουν 2026, 10_41_49 μ.μ."
   TextField "Text field_1" at 235,6 size 313x27; Text 'VFD PUMP PRESSURE CONTROL'
   TextField "Text field_2" at 335,42 size 128x25; Text 'DIAGNOSTICS'
   Button "Button_2" at 1,414 size 194x65; TextOff 'HOME'
      on Press: ActivateScreen("Main Overview", 0)
   Button "Button_3" at 195,414 size 204x65; TextOff 'CONTROL'
      on Press: ActivateScreen("Control", 0)
   Button "Button_4" at 398,414 size 200x65; TextOff 'ALARMS'
      on Press: ActivateScreen("Alarm Page", 0)
   Button "Button_5" at 597,414 size 200x65; TextOff 'DIAGNOSTICS'
      on Press: ActivateScreen("Diagnostics", 0)
   IOField "I/O field_2" at 44,352 size 50x27; FormatPattern 99.9
      ProcessValue <- "DB_VFD_Motor_Pressure_Actual"
   GraphicView "Graphic view_7" at 610,430 size 39x34; Picture "Graphic_1"
   GraphicView "Graphic view_8" at 422,429 size 43x33; Picture "Graphic_2"
   GraphicView "Graphic view_9" at 35,428 size 41x33; Picture "Graphic_3"
   GraphicView "Graphic view_10" at 213,430 size 36x30; Picture "Graphic_4"
   TextField "Text field_6" at 481,84 size 143x20; Text 'DIAGNOSTICS VALUES'
   Bar "Bar_1" at 47,127 size 45x212; MinimumValue 0; MaximumValue 100
      ProcessValue <- "DB_VFD_Motor_Pressure_Actual"
   Bar "Bar_2" at 145,127 size 45x212; MinimumValue 0; MaximumValue 100
      ProcessValue <- "DB_VFD_Motor_Pressure_Setpoint"
   Bar "Bar_3" at 244,127 size 45x212; MinimumValue 0; MaximumValue 100
      ProcessValue <- "DB_VFD_Motor_Actual_speed_hz"
   Bar "Bar_4" at 340,127 size 45x212; MinimumValue 0; MaximumValue 100
      ProcessValue <- "DB_VFD_Motor_Ramp_Output"
   IOField "I/O field_3" at 656,165 size 108x37; FormatPattern 99.9; Unit bar
      ProcessValue <- "DB_VFD_Motor_Max_Pressure_Limit"
   IOField "I/O field_4" at 664,210 size 100x37; FormatPattern 9.9; Unit Hz
      ProcessValue <- "DB_VFD_Motor_Ramp_Step"
   IOField "I/O field_5" at 656,255 size 108x37; FormatPattern 9999; Unit %
      ProcessValue <- "DB_VFD_Motor_Output_scaled"
   IOField "I/O field_6" at 640,300 size 124x37; FormatPattern 99.9; Unit bar
      ProcessValue <- "DB_VFD_Motor_Pressure_Actual"
   IOField "I/O field_7" at 664,346 size 100x37; FormatPattern 999
      ProcessValue <- "DB_VFD_Motor_Fault_code"
   TextField "Text field_3" at 482,127 size 136x20; Text 'MIN PRESSURE LIMIT'
   TextField "Text field_4" at 482,173 size 142x20; Text 'MAX PRESSURE LIMIT'
   TextField "Text field_5" at 483,221 size 77x20; Text 'RAMP STEP'
   TextField "Text field_7" at 483,264 size 105x20; Text 'OUTPUT SCALED'
   TextField "Text field_8" at 485,307 size 123x20; Text 'PRESSURE ACTUAL'
   TextField "Text field_9" at 485,352 size 80x20; Text 'FAULT CODE'
   TextField "Text field_10" at 34,75 size 69x52; Text 'ACTUAL PRESSURE (bar)'
   TextField "Text field_11" at 130,76 size 73x52; Text 'PRESSURE SETPOINT (bar)'
   TextField "Text field_12" at 239,76 size 59x52; Text 'ACTUAL SPEED (Hz)'
   TextField "Text field_13" at 336,75 size 56x52; Text 'RAMP OUTPUT (Hz)'
   IOField "I/O field_8" at 142,352 size 50x27; FormatPattern 99.9
      ProcessValue <- "DB_VFD_Motor_Pressure_Setpoint"
   IOField "I/O field_9" at 241,352 size 50x27; FormatPattern 99.9
      ProcessValue <- "DB_VFD_Motor_Actual_speed_hz"
   IOField "I/O field_10" at 338,352 size 50x27; FormatPattern 99.9
      ProcessValue <- "DB_VFD_Motor_Ramp_Output"
   IOField "I/O field_1" at 651,123 size 108x37; FormatPattern 99.9; Unit bar
      ProcessValue <- "DB_VFD_Motor_Min_Pressure_Limit"
*)